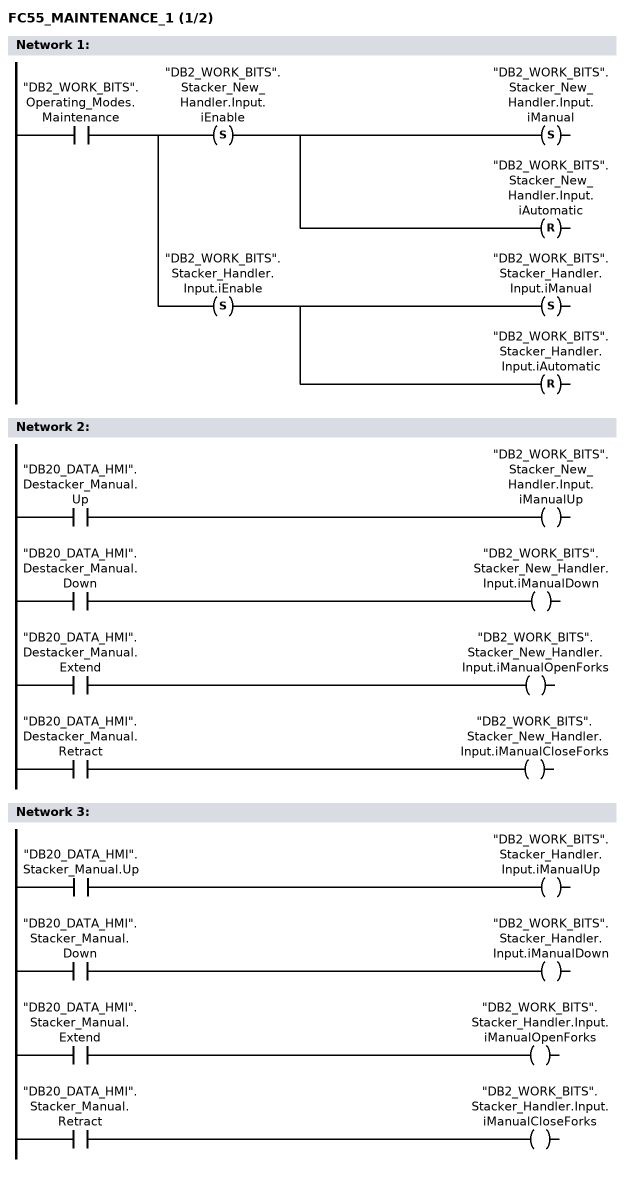
   RUNG wire#powerrail
      Contact( "DB2_WORK_BITS".Operating_Modes.Maintenance )
      wire#w1
      S_Coil( "DB2_WORK_BITS".Stacker_New_Handler.Input.iEnable )
      wire#w2
      S_Coil( "DB2_WORK_BITS".Stacker_New_Handler.Input.iManual )
   END_RUNG
   RUNG wire#w2
      R_Coil( "DB2_WORK_BITS".Stacker_New_Handler.Input.iAutomatic )
   END_RUNG
   RUNG wire#w1
      S_Coil( "DB2_WORK_BITS".Stacker_Handler.Input.iEnable )
      wire#w3
      S_Coil( "DB2_WORK_BITS".Stacker_Handler.Input.iManual )
   END_RUNG
   RUNG wire#w3
      R_Coil( "DB2_WORK_BITS".Stacker_Handler.Input.iAutomatic )
   END_RUNG
   // the same network as SCL:
   IF "DB2_WORK_BITS".Operating_Modes.Maintenance THEN
       "DB2_WORK_BITS".Stacker_New_Handler.Input.iEnable := TRUE;
       "DB2_WORK_BITS".Stacker_New_Handler.Input.iManual := TRUE;
       "DB2_WORK_BITS".Stacker_New_Handler.Input.iAutomatic := FALSE;
       "DB2_WORK_BITS".Stacker_Handler.Input.iEnable := TRUE;
       "DB2_WORK_BITS".Stacker_Handler.Input.iManual := TRUE;
       "DB2_WORK_BITS".Stacker_Handler.Input.iAutomatic := FALSE;
   END_IF;
END_REGION

REGION Network 2
   RUNG wire#powerrail
      Contact( "DB20_DATA_HMI".Destacker_Manual.Up )
      Coil( "DB2_WORK_BITS".Stacker_New_Handler.Input.iManualUp )
   END_RUNG
   RUNG wire#powerrail
      Contact( "DB20_DATA_HMI".Destacker_Manual.Down )
      Coil( "DB2_WORK_BITS".Stacker_New_Handler.Input.iManualDown )
   END_RUNG
   RUNG wire#powerrail
      Contact( "DB20_DATA_HMI".Destacker_Manual.Extend )
      Coil( "DB2_WORK_BITS".Stacker_New_Handler.Input.iManualOpenForks )
   END_RUNG
   RUNG wire#powerrail
      Contact( "DB20_DATA_HMI".Destacker_Manual.Retract )
      Coil( "DB2_WORK_BITS".Stacker_New_Handler.Input.iManualCloseForks )
   END_RUNG
   // the same network as SCL:
   "DB2_WORK_BITS".Stacker_New_Handler.Input.iManualUp := "DB20_DATA_HMI".Destacker_Manual.Up;
   "DB2_WORK_BITS".Stacker_New_Handler.Input.iManualDown := "DB20_DATA_HMI".Destacker_Manual.Down;
   "DB2_WORK_BITS".Stacker_New_Handler.Input.iManualOpenForks := "DB20_DATA_HMI".Destacker_Manual.Extend;
   "DB2_WORK_BITS".Stacker_New_Handler.Input.iManualCloseForks := "DB20_DATA_HMI".Destacker_Manual.Retract;
END_REGION

REGION Network 3
   RUNG wire#powerrail
      Contact( "DB20_DATA_HMI".Stacker_Manual.Up )
      Coil( "DB2_WORK_BITS".Stacker_Handler.Input.iManualUp )
   END_RUNG
   RUNG wire#powerrail
      Contact( "DB20_DATA_HMI".Stacker_Manual.Down )
      Coil( "DB2_WORK_BITS".Stacker_Handler.Input.iManualDown )
   END_RUNG
   RUNG wire#powerrail
      Contact( "DB20_DATA_HMI".Stacker_Manual.Extend )
      Coil( "DB2_WORK_BITS".Stacker_Handler.Input.iManualOpenForks )
   END_RUNG
   RUNG wire#powerrail
      Contact( "DB20_DATA_HMI".Stacker_Manual.Retract )
      Coil( "DB2_WORK_BITS".Stacker_Handler.Input.iManualCloseForks )
   END_RUNG
   // the same network as SCL:
   "DB2_WORK_BITS".Stacker_Handler.Input.iManualUp := "DB20_DATA_HMI".Stacker_Manual.Up;
   "DB2_WORK_BITS".Stacker_Handler.Input.iManualDown := "DB20_DATA_HMI".Stacker_Manual.Down;
   "DB2_WORK_BITS".Stacker_Handler.Input.iManualOpenForks := "DB20_DATA_HMI".Stacker_Manual.Extend;
   "DB2_WORK_BITS".Stacker_Handler.Input.iManualCloseForks := "DB20_DATA_HMI".Stacker_Manual.Retract;
END_REGION

REGION Network 4
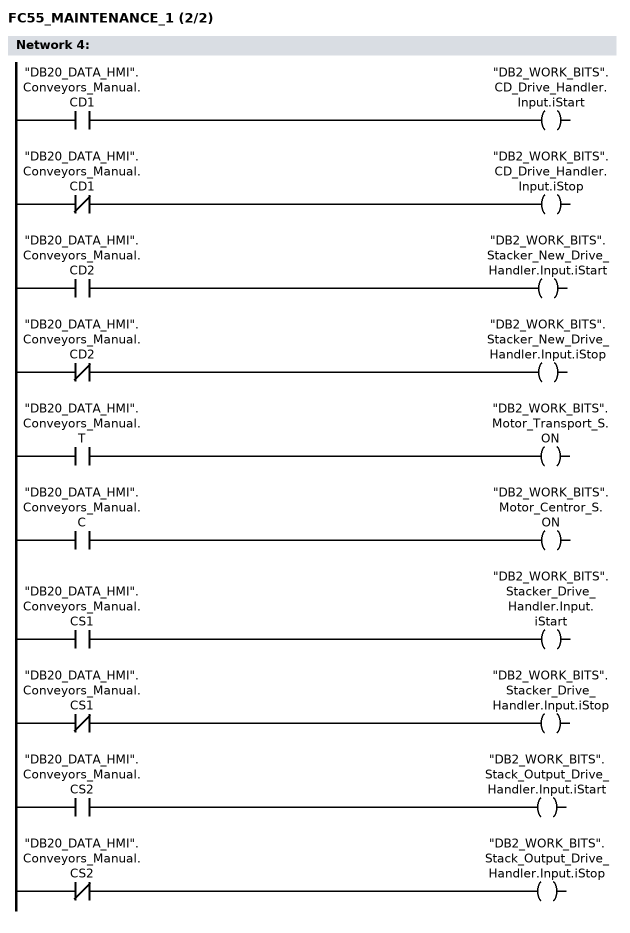
   RUNG wire#powerrail
      Contact( "DB20_DATA_HMI".Conveyors_Manual.CD1 )
      Coil( "DB2_WORK_BITS".CD_Drive_Handler.Input.iStart )
   END_RUNG
   RUNG wire#powerrail
      I_Contact( "DB20_DATA_HMI".Conveyors_Manual.CD1 )
      Coil( "DB2_WORK_BITS".CD_Drive_Handler.Input.iStop )
   END_RUNG
   RUNG wire#powerrail
      Contact( "DB20_DATA_HMI".Conveyors_Manual.CD2 )
      Coil( "DB2_WORK_BITS".Stacker_New_Drive_Handler.Input.iStart )
   END_RUNG
   RUNG wire#powerrail
      I_Contact( "DB20_DATA_HMI".Conveyors_Manual.CD2 )
      Coil( "DB2_WORK_BITS".Stacker_New_Drive_Handler.Input.iStop )
   END_RUNG
   RUNG wire#powerrail
      Contact( "DB20_DATA_HMI".Conveyors_Manual.T )
      Coil( "DB2_WORK_BITS".Motor_Transport_S.ON )
   END_RUNG
   RUNG wire#powerrail
      Contact( "DB20_DATA_HMI".Conveyors_Manual.C )
      Coil( "DB2_WORK_BITS".Motor_Centror_S.ON )
   END_RUNG
   RUNG wire#powerrail
      Contact( "DB20_DATA_HMI".Conveyors_Manual.CS1 )
      Coil( "DB2_WORK_BITS".Stacker_Drive_Handler.Input.iStart )
   END_RUNG
   RUNG wire#powerrail
      I_Contact( "DB20_DATA_HMI".Conveyors_Manual.CS1 )
      Coil( "DB2_WORK_BITS".Stacker_Drive_Handler.Input.iStop )
   END_RUNG
   RUNG wire#powerrail
      Contact( "DB20_DATA_HMI".Conveyors_Manual.CS2 )
      Coil( "DB2_WORK_BITS".Stack_Output_Drive_Handler.Input.iStart )
   END_RUNG
   RUNG wire#powerrail
      I_Contact( "DB20_DATA_HMI".Conveyors_Manual.CS2 )
      Coil( "DB2_WORK_BITS".Stack_Output_Drive_Handler.Input.iStop )
   END_RUNG
   // the same network as SCL:
   "DB2_WORK_BITS".CD_Drive_Handler.Input.iStart := "DB20_DATA_HMI".Conveyors_Manual.CD1;
   "DB2_WORK_BITS".CD_Drive_Handler.Input.iStop := NOT "DB20_DATA_HMI".Conveyors_Manual.CD1;
   "DB2_WORK_BITS".Stacker_New_Drive_Handler.Input.iStart := "DB20_DATA_HMI".Conveyors_Manual.CD2;
   "DB2_WORK_BITS".Stacker_New_Drive_Handler.Input.iStop := NOT "DB20_DATA_HMI".Conveyors_Manual.CD2;
   "DB2_WORK_BITS".Motor_Transport_S.ON := "DB20_DATA_HMI".Conveyors_Manual.T;
   "DB2_WORK_BITS".Motor_Centror_S.ON := "DB20_DATA_HMI".Conveyors_Manual.C;
   "DB2_WORK_BITS".Stacker_Drive_Handler.Input.iStart := "DB20_DATA_HMI".Conveyors_Manual.CS1;
   "DB2_WORK_BITS".Stacker_Drive_Handler.Input.iStop := NOT "DB20_DATA_HMI".Conveyors_Manual.CS1;
   "DB2_WORK_BITS".Stack_Output_Drive_Handler.Input.iStart := "DB20_DATA_HMI".Conveyors_Manual.CS2;
   "DB2_WORK_BITS".Stack_Output_Drive_Handler.Input.iStop := NOT "DB20_DATA_HMI".Conveyors_Manual.CS2;
END_REGION
END_FUNCTION

FUNCTION "FC58_SAFETY" : Void   // FC58, LAD
{ S7_Optimized_Access := 'TRUE' }
VERSION : 0.1
BEGIN

REGION Network 1: Stacker
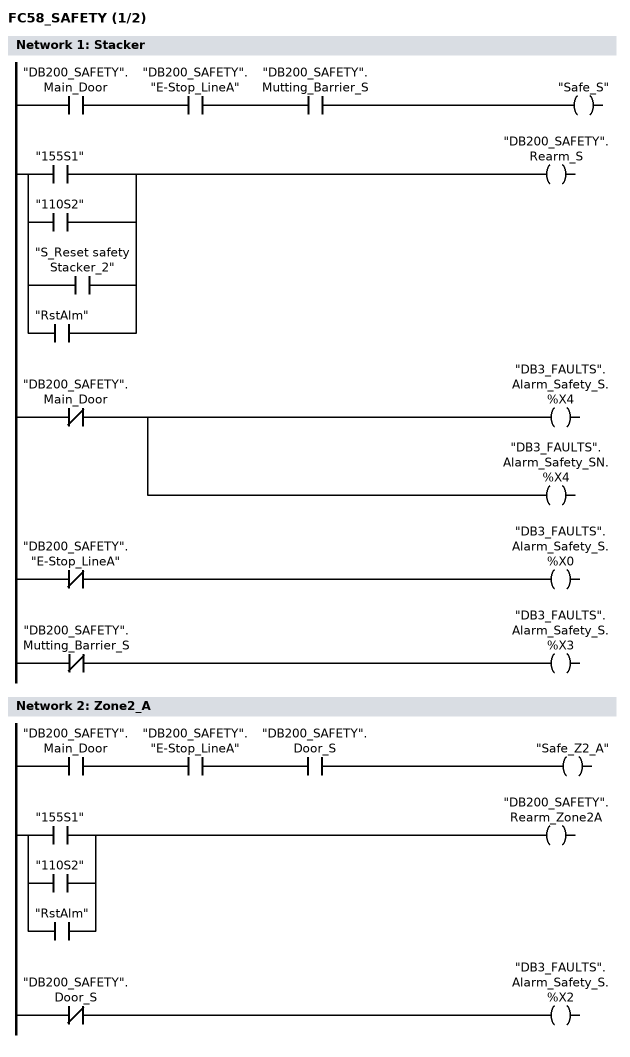
   RUNG wire#powerrail
      Contact( "DB200_SAFETY".Main_Door )
      Contact( "DB200_SAFETY"."E-Stop_LineA" )
      Contact( "DB200_SAFETY".Mutting_Barrier_S )
      Coil( "Safe_S" )
   END_RUNG
   RUNG wire#powerrail
      Contact( "155S1" )
      wire#w1
      Coil( "DB200_SAFETY".Rearm_S )
   END_RUNG
   RUNG wire#powerrail
      Contact( "110S2" )
   END_RUNG wire#w1
   RUNG wire#powerrail
      Contact( "S_Reset safety Stacker_2" )
   END_RUNG wire#w1
   RUNG wire#powerrail
      Contact( "RstAlm" )
   END_RUNG wire#w1
   RUNG wire#powerrail
      I_Contact( "DB200_SAFETY".Main_Door )
      wire#w2
      Coil( "DB3_FAULTS".Alarm_Safety_S.%X4 )
   END_RUNG
   RUNG wire#w2
      Coil( "DB3_FAULTS".Alarm_Safety_SN.%X4 )
   END_RUNG
   RUNG wire#powerrail
      I_Contact( "DB200_SAFETY"."E-Stop_LineA" )
      Coil( "DB3_FAULTS".Alarm_Safety_S.%X0 )
   END_RUNG
   RUNG wire#powerrail
      I_Contact( "DB200_SAFETY".Mutting_Barrier_S )
      Coil( "DB3_FAULTS".Alarm_Safety_S.%X3 )
   END_RUNG
   // the same network as SCL:
   "Safe_S" := "DB200_SAFETY".Main_Door AND "DB200_SAFETY"."E-Stop_LineA" AND "DB200_SAFETY".Mutting_Barrier_S;
   "DB200_SAFETY".Rearm_S := "155S1" OR "110S2" OR "S_Reset safety Stacker_2" OR "RstAlm";
   "DB3_FAULTS".Alarm_Safety_S.%X4 := NOT "DB200_SAFETY".Main_Door;
   "DB3_FAULTS".Alarm_Safety_SN.%X4 := NOT "DB200_SAFETY".Main_Door;
   "DB3_FAULTS".Alarm_Safety_S.%X0 := NOT "DB200_SAFETY"."E-Stop_LineA";
   "DB3_FAULTS".Alarm_Safety_S.%X3 := NOT "DB200_SAFETY".Mutting_Barrier_S;
END_REGION

REGION Network 2: Zone2_A
   RUNG wire#powerrail
      Contact( "DB200_SAFETY".Main_Door )
      Contact( "DB200_SAFETY"."E-Stop_LineA" )
      Contact( "DB200_SAFETY".Door_S )
      Coil( "Safe_Z2_A" )
   END_RUNG
   RUNG wire#powerrail
      Contact( "155S1" )
      wire#w1
      Coil( "DB200_SAFETY".Rearm_Zone2A )
   END_RUNG
   RUNG wire#powerrail
      Contact( "110S2" )
   END_RUNG wire#w1
   RUNG wire#powerrail
      Contact( "RstAlm" )
   END_RUNG wire#w1
   RUNG wire#powerrail
      I_Contact( "DB200_SAFETY".Door_S )
      Coil( "DB3_FAULTS".Alarm_Safety_S.%X2 )
   END_RUNG
   // the same network as SCL:
   "Safe_Z2_A" := "DB200_SAFETY".Main_Door AND "DB200_SAFETY"."E-Stop_LineA" AND "DB200_SAFETY".Door_S;
   "DB200_SAFETY".Rearm_Zone2A := "155S1" OR "110S2" OR "RstAlm";
   "DB3_FAULTS".Alarm_Safety_S.%X2 := NOT "DB200_SAFETY".Door_S;
END_REGION

REGION Network 3: Stacker_New
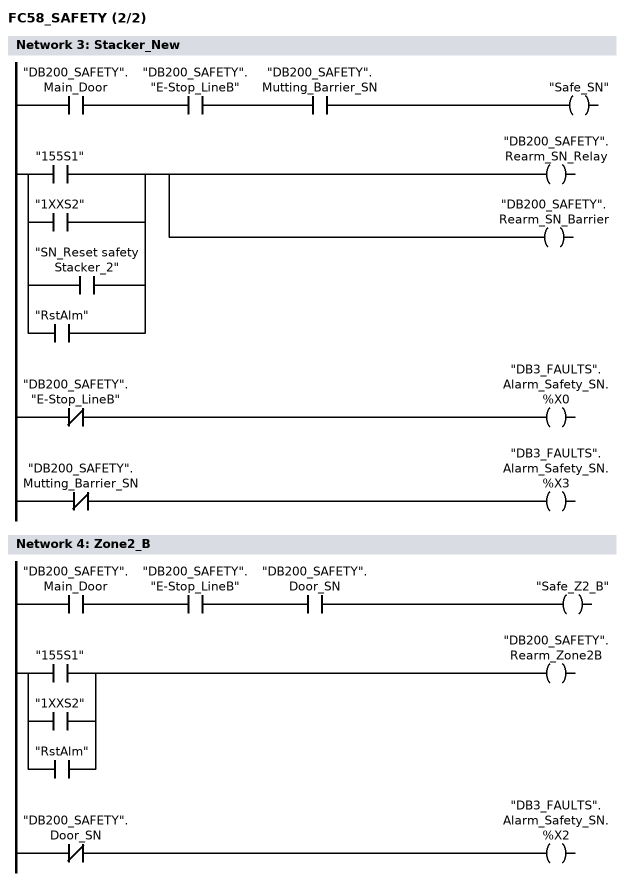
   RUNG wire#powerrail
      Contact( "DB200_SAFETY".Main_Door )
      Contact( "DB200_SAFETY"."E-Stop_LineB" )
      Contact( "DB200_SAFETY".Mutting_Barrier_SN )
      Coil( "Safe_SN" )
   END_RUNG
   RUNG wire#powerrail
      Contact( "155S1" )
      wire#w1
      Coil( "DB200_SAFETY".Rearm_SN_Relay )
   END_RUNG
   RUNG wire#powerrail
      Contact( "1XXS2" )
   END_RUNG wire#w1
   RUNG wire#powerrail
      Contact( "SN_Reset safety Stacker_2" )
   END_RUNG wire#w1
   RUNG wire#powerrail
      Contact( "RstAlm" )
   END_RUNG wire#w1
   RUNG wire#w1
      Coil( "DB200_SAFETY".Rearm_SN_Barrier )
   END_RUNG
   RUNG wire#powerrail
      I_Contact( "DB200_SAFETY"."E-Stop_LineB" )
      Coil( "DB3_FAULTS".Alarm_Safety_SN.%X0 )
   END_RUNG
   RUNG wire#powerrail
      I_Contact( "DB200_SAFETY".Mutting_Barrier_SN )
      Coil( "DB3_FAULTS".Alarm_Safety_SN.%X3 )
   END_RUNG
   // the same network as SCL:
   "Safe_SN" := "DB200_SAFETY".Main_Door AND "DB200_SAFETY"."E-Stop_LineB" AND "DB200_SAFETY".Mutting_Barrier_SN;
   "DB200_SAFETY".Rearm_SN_Relay := "155S1" OR "1XXS2" OR "SN_Reset safety Stacker_2" OR "RstAlm";
   "DB200_SAFETY".Rearm_SN_Barrier := "DB200_SAFETY".Rearm_SN_Relay;
   "DB3_FAULTS".Alarm_Safety_SN.%X0 := NOT "DB200_SAFETY"."E-Stop_LineB";
   "DB3_FAULTS".Alarm_Safety_SN.%X3 := NOT "DB200_SAFETY".Mutting_Barrier_SN;
END_REGION

REGION Network 4: Zone2_B
   RUNG wire#powerrail
      Contact( "DB200_SAFETY".Main_Door )
      Contact( "DB200_SAFETY"."E-Stop_LineB" )
      Contact( "DB200_SAFETY".Door_SN )
      Coil( "Safe_Z2_B" )
   END_RUNG
   RUNG wire#powerrail
      Contact( "155S1" )
      wire#w1
      Coil( "DB200_SAFETY".Rearm_Zone2B )
   END_RUNG
   RUNG wire#powerrail
      Contact( "1XXS2" )
   END_RUNG wire#w1
   RUNG wire#powerrail
      Contact( "RstAlm" )
   END_RUNG wire#w1
   RUNG wire#powerrail
      I_Contact( "DB200_SAFETY".Door_SN )
      Coil( "DB3_FAULTS".Alarm_Safety_SN.%X2 )
   END_RUNG
   // the same network as SCL:
   "Safe_Z2_B" := "DB200_SAFETY".Main_Door AND "DB200_SAFETY"."E-Stop_LineB" AND "DB200_SAFETY".Door_SN;
   "DB200_SAFETY".Rearm_Zone2B := "155S1" OR "1XXS2" OR "RstAlm";
   "DB3_FAULTS".Alarm_Safety_SN.%X2 := NOT "DB200_SAFETY".Door_SN;
END_REGION
END_FUNCTION

FUNCTION "FC100_CountDaily" : Void   // FC100, SCL
{ S7_Optimized_Access := 'TRUE' }
VERSION : 0.1
   VAR_INPUT
      SignalToCount : Bool;
      Reset : Bool;
   END_VAR
   VAR_IN_OUT
      CurrentValue : UDInt;
   END_VAR
   VAR_TEMP
      timeofday : DTL;
      ret : Int;
   END_VAR
BEGIN
   #ret := RD_LOC_T(#timeofday);
END_FUNCTION

ORGANIZATION_BLOCK "Main"   // OB1, LAD, ProgramCycle
TITLE = "Main Program Sweep (Cycle)"
{ S7_Optimized_Access := 'TRUE' }
VERSION : 0.1
   VAR_INPUT
      Initial_Call : Bool;   // Initial call of this OB
      Remanence : Bool;   // =True, if remanent data are available
   END_VAR
   VAR_TEMP
      Move_Block_Diag : Int;
   END_VAR
BEGIN

REGION Network 1
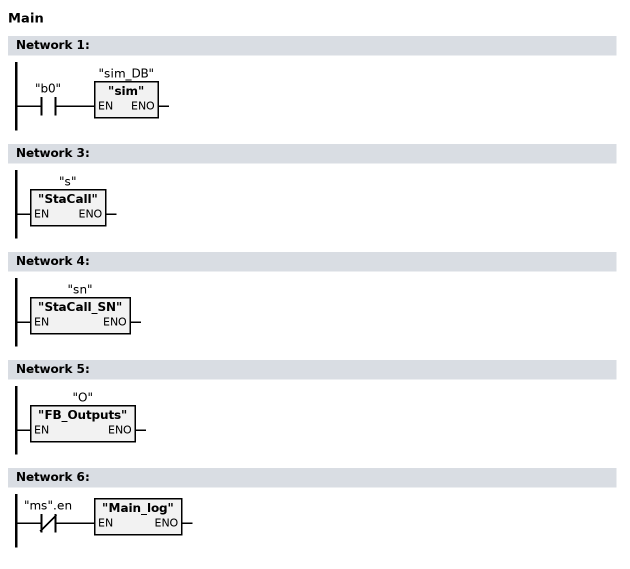
   RUNG wire#powerrail
      Contact( "b0" )
      "sim_DB"()
   END_RUNG
   // the same network as SCL:
   IF "b0" THEN
       "sim_DB"();   // "sim"
   END_IF;
END_REGION

REGION Network 2 (SCL)
   "FC58_SAFETY"();
   "FC6_OUTPUTS"();

   "FC60_MappingIn"();

   "FC3_FAULTS"();
   "FB_GEN_DB"();

   "FC_AckOpTranzit"();


   "FC52_STACKING"();
   "FC52_STACKING_New"();

   //"FC55_MAINTENANCE"();
   "FC20_HMI"();
   "FB_IntervalTrigger_DB"();
   "FB_EnergyCounter_DB"(ibMeterPulse := "DB2_WORK_BITS".Consumption_Pulse,
                         ibHourChange := "FB_IntervalTrigger_DB".bHourChanged,
                        ibDayChange := "FB_IntervalTrigger_DB".bDayChanged,
                         ibMonthChange := "FB_IntervalTrigger_DB".bMonthChanged,
                         ibReset := FALSE);
   "FB_AlarmCounter_DB"();
   "FB_ProductionStatistics_DB"(ibDestroy:="DB2_WORK_BITS".SQ_Outfeed_Stack_SN,
                                ibRepair:="DB2_WORK_BITS".Transport_Conveyor_SQs.SQ_Repaired_Pallet[0] OR "DB2_WORK_BITS".Transport_Conveyor_SQs.SQ_Repaired_Pallet[1],
                                ibDayChange:="FB_IntervalTrigger_DB".bDayChanged,
                                ibMonthChange:="FB_IntervalTrigger_DB".bMonthChanged);
END_REGION

REGION Network 3
   RUNG wire#powerrail
      "s"()
   END_RUNG
   // the same network as SCL:
   "s"();   // "StaCall"
END_REGION

REGION Network 4
   RUNG wire#powerrail
      "sn"()
   END_RUNG
   // the same network as SCL:
   "sn"();   // "StaCall_SN"
END_REGION

REGION Network 5
   RUNG wire#powerrail
      "O"()
   END_RUNG
   // the same network as SCL:
   "O"();   // "FB_Outputs"
END_REGION

REGION Network 6
   RUNG wire#powerrail
      I_Contact( "ms".en )
      "Main_log"()
   END_RUNG
   // the same network as SCL:
   IF NOT "ms".en THEN "Main_log"(); END_IF;
END_REGION
END_ORGANIZATION_BLOCK

ORGANIZATION_BLOCK "OB82_I/O_FLT"   // OB82, LAD, DiagnosticErrorInterrupt
{ S7_Optimized_Access := 'TRUE' }
VERSION : 0.1
   VAR_INPUT
      IO_State : Word;   // IO state of the HW object
      LADDR : Hw_Any;   // Hardware identifier
      Channel : UInt;   // Channel number
      MultiError : Bool;   // =true if more than one error is present
   END_VAR
BEGIN
END_ORGANIZATION_BLOCK

ORGANIZATION_BLOCK "OB100_COMPLETE_RESTART"   // OB100, LAD, Startup
TITLE = "Complete Restart"
{ S7_Optimized_Access := 'TRUE' }
VERSION : 0.1
   VAR_INPUT
      LostRetentive : Bool;   // True if retentive data are lost
      LostRTC : Bool;   // True if date and time are lost
   END_VAR
BEGIN
END_ORGANIZATION_BLOCK

// folder: Stacker_New

FUNCTION_BLOCK "StaCall_SN"   // FB15, LAD
{ S7_Optimized_Access := 'TRUE' }
VERSION : 0.1
   VAR
      f : Array[0..10] of "sta_SN";
      tranzit : Array[0..10] of Bool;
      Range_LS_1 : Bool;
      Range_LS_2 : Bool;
      Range_LS_3 : Bool;
      PrezPalStackLength : Bool;
      PrezPalStackAnyLength : Bool;
      PrezPalStackAny : Bool;
      DeliveryStack : Bool;
      StivStat : USInt;
      nAc : USInt;
      tmrSnzCentr : TON_TIME;
      tmr : Array[0..8] of IEC_TIMER;
   END_VAR
   VAR_TEMP
      to_ce : Bool;
      to_cm : Bool;
      cmdLiftUpO : Bool;
      tranzit12 : Bool;
   END_VAR
   VAR CONSTANT
      _nop0 : Int := 0;
      _op1 : Int := 1;
      _cen : Int := 3;
      _stack : Int := 4;
      _evac : Int := 5;
      _nop : Int := 6;
   END_VAR
   VAR_TEMP   // added for the SCL form of the ladder/FBD networks
      _w1 : Bool;
      _w2 : Bool;
      _w3 : Bool;
   END_VAR
BEGIN

REGION Network 1: Force init
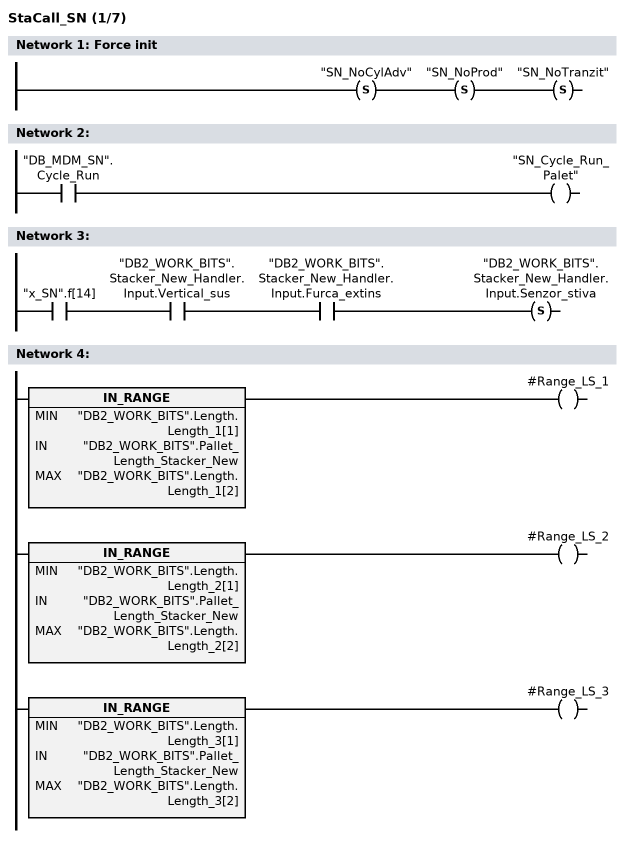
   RUNG wire#powerrail
      S_Coil( "SN_NoCylAdv" )
      S_Coil( "SN_NoProd" )
      S_Coil( "SN_NoTranzit" )
   END_RUNG
   // the same network as SCL:
   "SN_NoCylAdv" := TRUE;
   "SN_NoProd" := TRUE;
   "SN_NoTranzit" := TRUE;
END_REGION

REGION Network 2
   RUNG wire#powerrail
      Contact( "DB_MDM_SN".Cycle_Run )
      Coil( "SN_Cycle_Run_Palet" )
   END_RUNG
   // the same network as SCL:
   "SN_Cycle_Run_Palet" := "DB_MDM_SN".Cycle_Run;
END_REGION

REGION Network 3
   RUNG wire#powerrail
      Contact( "x_SN".f[14] )
      Contact( "DB2_WORK_BITS".Stacker_New_Handler.Input.Vertical_sus )
      Contact( "DB2_WORK_BITS".Stacker_New_Handler.Input.Furca_extins )
      S_Coil( "DB2_WORK_BITS".Stacker_New_Handler.Input.Senzor_stiva )
   END_RUNG
   // the same network as SCL:
   IF "x_SN".f[14] AND "DB2_WORK_BITS".Stacker_New_Handler.Input.Vertical_sus AND "DB2_WORK_BITS".Stacker_New_Handler.Input.Furca_extins THEN
       "DB2_WORK_BITS".Stacker_New_Handler.Input.Senzor_stiva := TRUE;
   END_IF;
END_REGION

REGION Network 4
   RUNG wire#powerrail
      { S7_Templates := "SrcType := Int" } InRange(min := "DB2_WORK_BITS".Length.Length_1[1], in := "DB2_WORK_BITS".Pallet_Length_Stacker_New, max := "DB2_WORK_BITS".Length.Length_1[2])
      Coil( #Range_LS_1 )
   END_RUNG
   RUNG wire#powerrail
      { S7_Templates := "SrcType := Int" } InRange(min := "DB2_WORK_BITS".Length.Length_2[1], in := "DB2_WORK_BITS".Pallet_Length_Stacker_New, max := "DB2_WORK_BITS".Length.Length_2[2])
      Coil( #Range_LS_2 )
   END_RUNG
   RUNG wire#powerrail
      { S7_Templates := "SrcType := Int" } InRange(min := "DB2_WORK_BITS".Length.Length_3[1], in := "DB2_WORK_BITS".Pallet_Length_Stacker_New, max := "DB2_WORK_BITS".Length.Length_3[2])
      Coil( #Range_LS_3 )
   END_RUNG
   // the same network as SCL:
   #Range_LS_1 := ("DB2_WORK_BITS".Length.Length_1[1] <= "DB2_WORK_BITS".Pallet_Length_Stacker_New) AND ("DB2_WORK_BITS".Pallet_Length_Stacker_New <= "DB2_WORK_BITS".Length.Length_1[2]);
   #Range_LS_2 := ("DB2_WORK_BITS".Length.Length_2[1] <= "DB2_WORK_BITS".Pallet_Length_Stacker_New) AND ("DB2_WORK_BITS".Pallet_Length_Stacker_New <= "DB2_WORK_BITS".Length.Length_2[2]);
   #Range_LS_3 := ("DB2_WORK_BITS".Length.Length_3[1] <= "DB2_WORK_BITS".Pallet_Length_Stacker_New) AND ("DB2_WORK_BITS".Pallet_Length_Stacker_New <= "DB2_WORK_BITS".Length.Length_3[2]);
END_REGION

REGION Network 5: 1 Op1- - Reparare palete Zona B
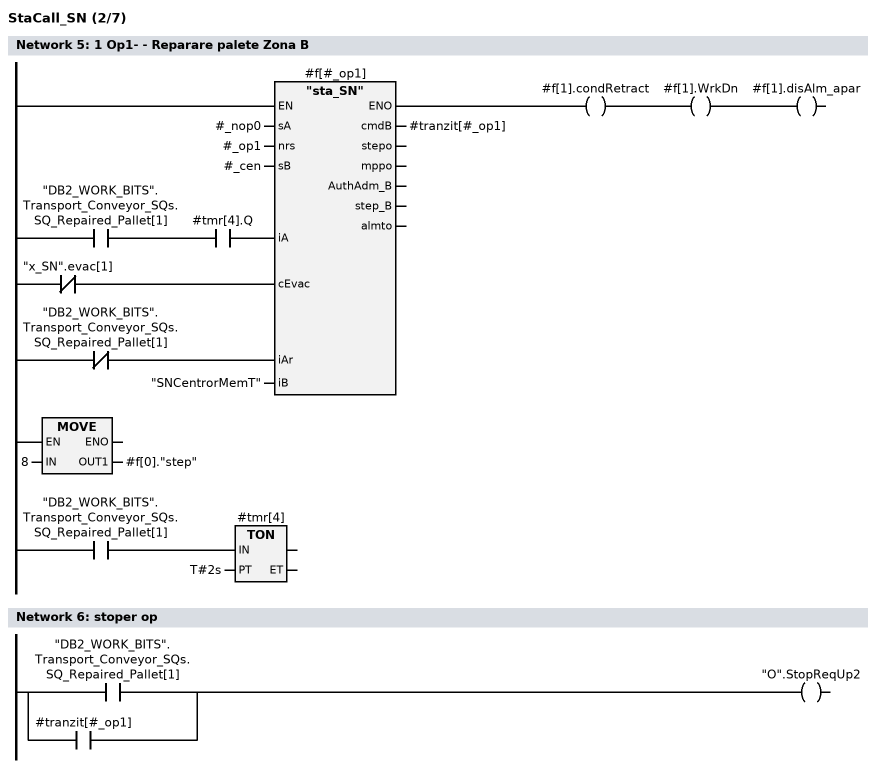
   #f[#_op1](sA := #_nop0,   // "sta_SN"
             nrs := #_op1,
             sB := #_cen,
             iA := "DB2_WORK_BITS".Transport_Conveyor_SQs.SQ_Repaired_Pallet[1] AND #tmr[4].Q,
             cEvac := NOT "x_SN".evac[1],
             iAr := NOT "DB2_WORK_BITS".Transport_Conveyor_SQs.SQ_Repaired_Pallet[1],
             iB := "SNCentrorMemT",
             cmdB => #tranzit[#_op1],
             ENO => #_w1);
   #f[1].condRetract := #_w1;
   #f[1].WrkDn := #_w1;
   #f[1].disAlm_apar := #_w1;
   #f[0]."step" := 8;
   #tmr[4].TON(IN := "DB2_WORK_BITS".Transport_Conveyor_SQs.SQ_Repaired_Pallet[1], PT := T#2s);
END_REGION

REGION Network 6: stoper op
   RUNG wire#powerrail
      Contact( "DB2_WORK_BITS".Transport_Conveyor_SQs.SQ_Repaired_Pallet[1] )
      wire#w1
      Coil( "O".StopReqUp2 )
   END_RUNG
   RUNG wire#powerrail
      Contact( #tranzit[#_op1] )
   END_RUNG wire#w1
   // the same network as SCL:
   "O".StopReqUp2 := "DB2_WORK_BITS".Transport_Conveyor_SQs.SQ_Repaired_Pallet[1] OR #tranzit[#_op1];
END_REGION

REGION Network 7
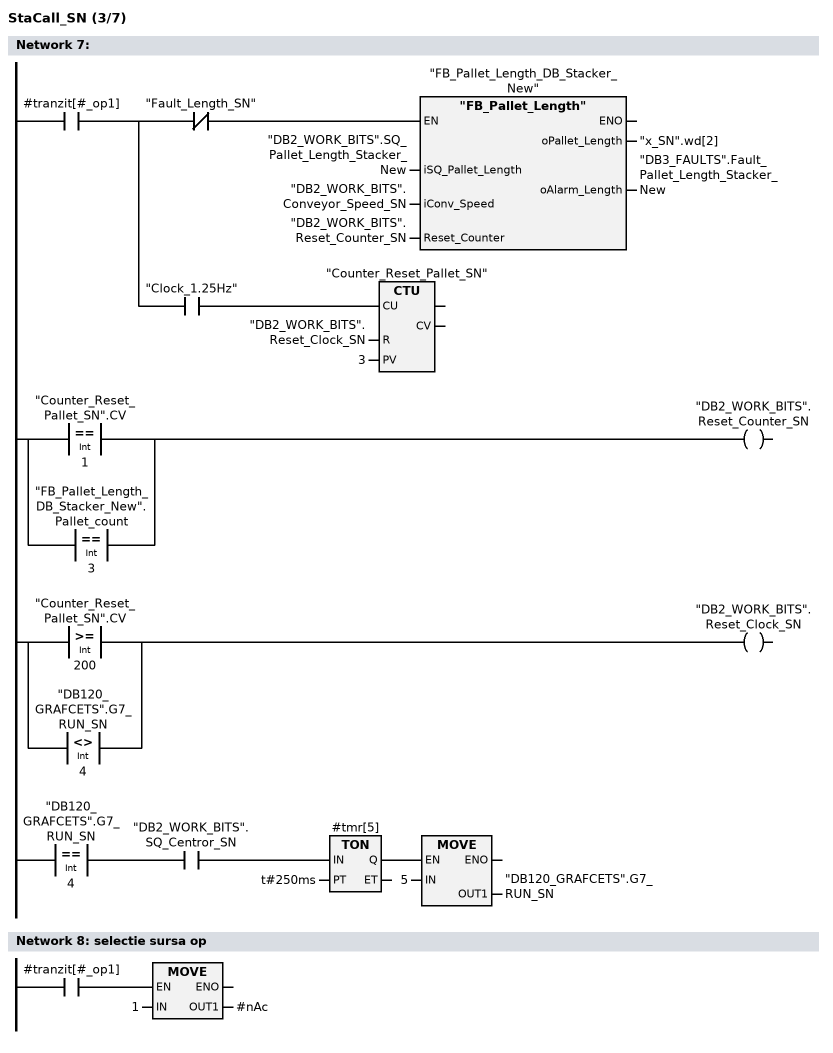
   IF #tranzit[#_op1] AND NOT "Fault_Length_SN" THEN
       "FB_Pallet_Length_DB_Stacker_New"(iSQ_Pallet_Length := "DB2_WORK_BITS".SQ_Pallet_Length_Stacker_New,   // "FB_Pallet_Length"
                               iConv_Speed := "DB2_WORK_BITS".Conveyor_Speed_SN,
                               Reset_Counter := "DB2_WORK_BITS".Reset_Counter_SN,
                               oPallet_Length => "x_SN".wd[2],
                               oAlarm_Length => "DB3_FAULTS".Fault_Pallet_Length_Stacker_New);
   END_IF;
   "Counter_Reset_Pallet_SN".CTU(CU := #tranzit[#_op1] AND "Clock_1.25Hz",
                           R := "DB2_WORK_BITS".Reset_Clock_SN,
                           PV := 3);
   "DB2_WORK_BITS".Reset_Counter_SN := ("Counter_Reset_Pallet_SN".CV = 1) OR ("FB_Pallet_Length_DB_Stacker_New".Pallet_count = 3);
   "DB2_WORK_BITS".Reset_Clock_SN := ("Counter_Reset_Pallet_SN".CV >= 200) OR ("DB120_GRAFCETS".G7_RUN_SN <> 4);
   #tmr[5].TON(IN := ("DB120_GRAFCETS".G7_RUN_SN = 4) AND "DB2_WORK_BITS".SQ_Centror_SN, PT := t#250ms);
   IF #tmr[5].Q THEN "DB120_GRAFCETS".G7_RUN_SN := 5; END_IF;
END_REGION

REGION Network 8: selectie sursa op
   RUNG wire#powerrail
      Contact( #tranzit[#_op1] )
      Move(in := 1, out1 => #nAc)
   END_RUNG
   // the same network as SCL:
   IF #tranzit[#_op1] THEN #nAc := 1; END_IF;
END_REGION

REGION Network 9: senz stop stk
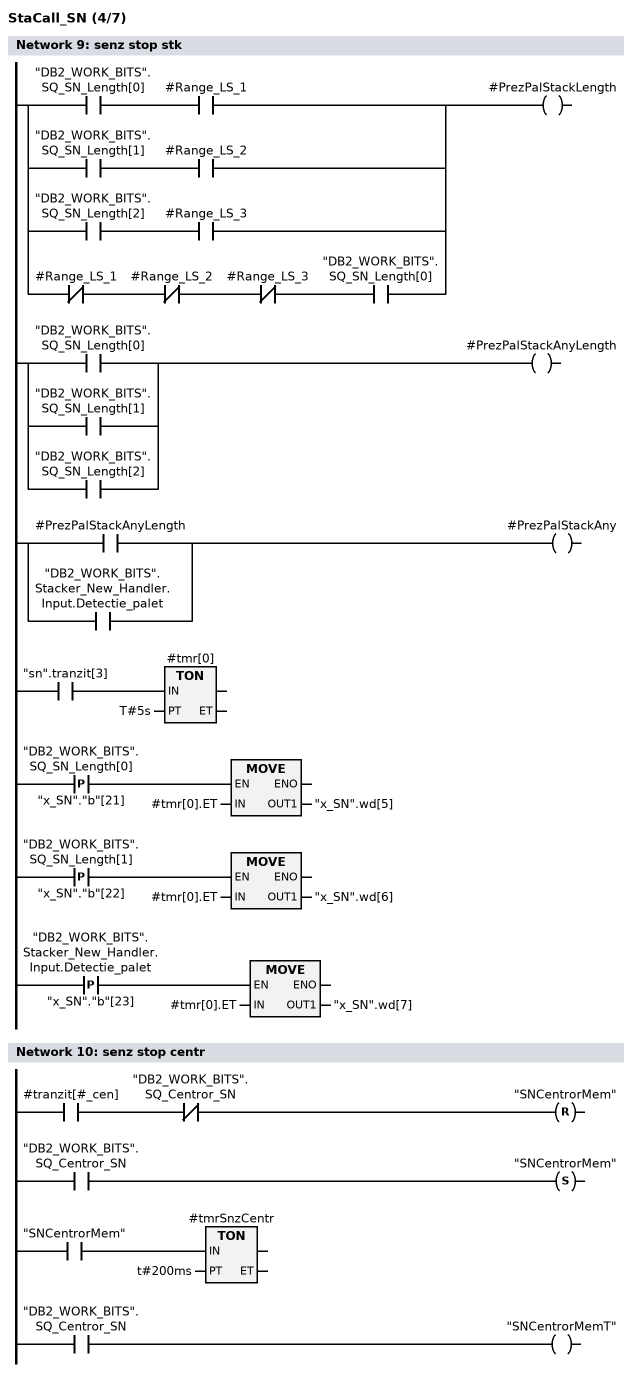
   #PrezPalStackLength := ("DB2_WORK_BITS".SQ_SN_Length[0] AND #Range_LS_1) OR ("DB2_WORK_BITS".SQ_SN_Length[1] AND #Range_LS_2) OR ("DB2_WORK_BITS".SQ_SN_Length[2] AND #Range_LS_3) OR (NOT #Range_LS_1 AND NOT #Range_LS_2 AND NOT #Range_LS_3 AND "DB2_WORK_BITS".SQ_SN_Length[0]);
   #PrezPalStackAnyLength := "DB2_WORK_BITS".SQ_SN_Length[0] OR "DB2_WORK_BITS".SQ_SN_Length[1] OR "DB2_WORK_BITS".SQ_SN_Length[2];
   #PrezPalStackAny := #PrezPalStackAnyLength OR "DB2_WORK_BITS".Stacker_New_Handler.Input.Detectie_palet;
   #tmr[0].TON(IN := "sn".tranzit[3], PT := T#5s);
   #_w1 := "DB2_WORK_BITS".SQ_SN_Length[0] AND NOT "x_SN"."b"[21];   // rising edge of "DB2_WORK_BITS".SQ_SN_Length[0]
   "x_SN"."b"[21] := "DB2_WORK_BITS".SQ_SN_Length[0];
   IF #_w1 THEN "x_SN".wd[5] := #tmr[0].ET; END_IF;
   #_w2 := "DB2_WORK_BITS".SQ_SN_Length[1] AND NOT "x_SN"."b"[22];   // rising edge of "DB2_WORK_BITS".SQ_SN_Length[1]
   "x_SN"."b"[22] := "DB2_WORK_BITS".SQ_SN_Length[1];
   IF #_w2 THEN "x_SN".wd[6] := #tmr[0].ET; END_IF;
   #_w3 := "DB2_WORK_BITS".Stacker_New_Handler.Input.Detectie_palet AND NOT "x_SN"."b"[23];   // rising edge of "DB2_WORK_BITS".Stacker_New_Handler.Input.Detectie_palet
   "x_SN"."b"[23] := "DB2_WORK_BITS".Stacker_New_Handler.Input.Detectie_palet;
   IF #_w3 THEN "x_SN".wd[7] := #tmr[0].ET; END_IF;
END_REGION

REGION Network 10: senz stop centr
   IF #tranzit[#_cen] AND NOT "DB2_WORK_BITS".SQ_Centror_SN THEN "SNCentrorMem" := FALSE; END_IF;
   IF "DB2_WORK_BITS".SQ_Centror_SN THEN "SNCentrorMem" := TRUE; END_IF;
   #tmrSnzCentr(IN := "SNCentrorMem", PT := t#200ms);   // TON
   "SNCentrorMemT" := "DB2_WORK_BITS".SQ_Centror_SN;
END_REGION

REGION Network 11: 3- Centror
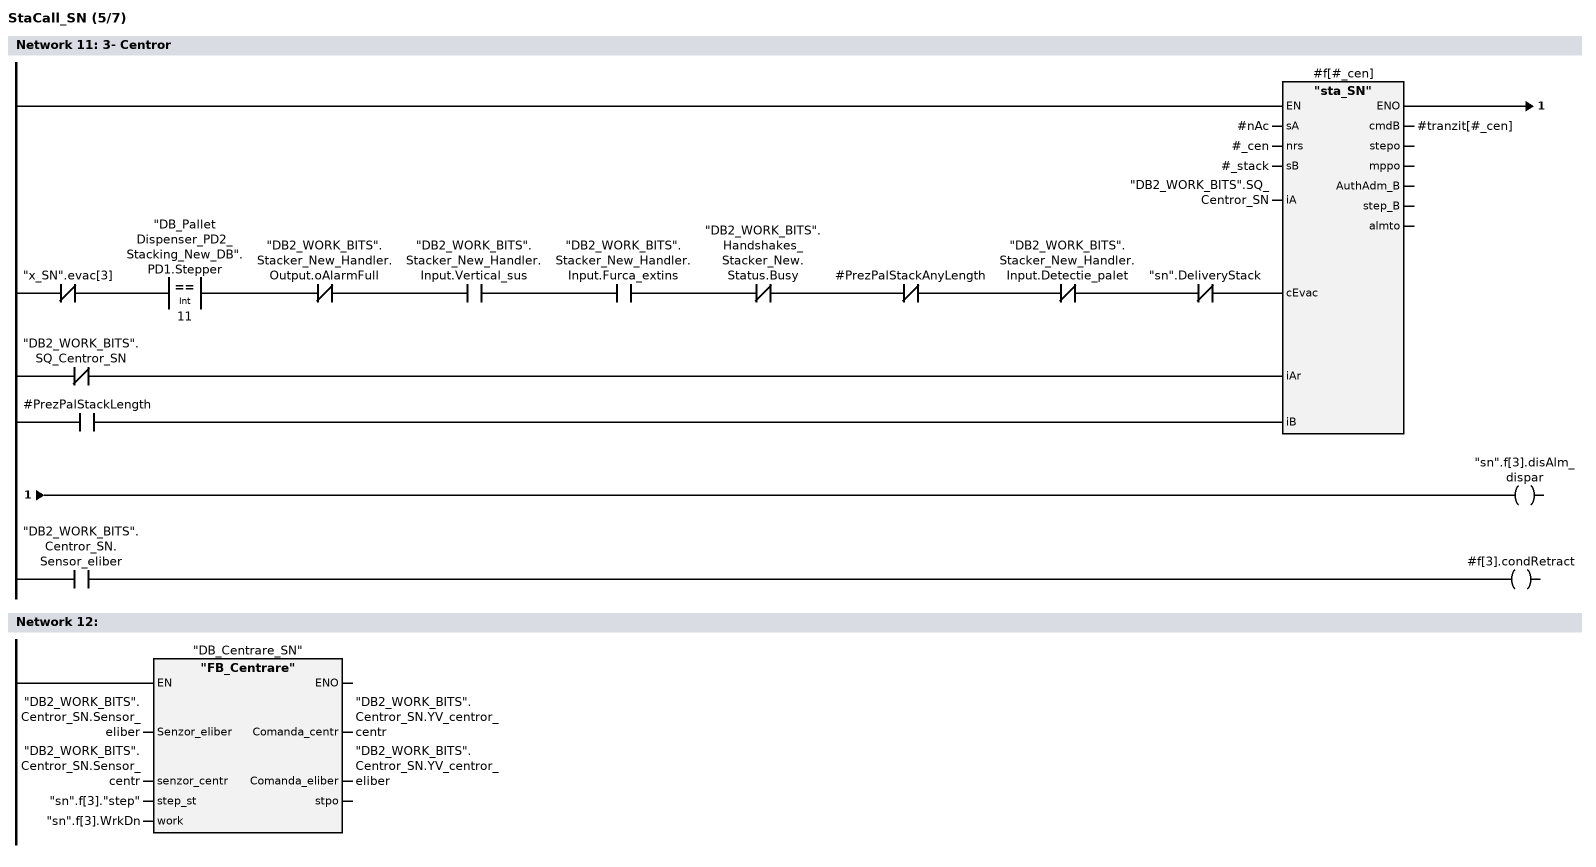
   RUNG wire#powerrail
      #f[#_cen](cEvac := wire#w1, iAr := wire#w2, iB := wire#w3, sA := #nAc, nrs := #_cen, sB := #_stack, iA := "DB2_WORK_BITS".SQ_Centror_SN, cmdB => #tranzit[#_cen], stepo =>, mppo =>, AuthAdm_B =>, step_B =>, almto =>)
      Coil( "sn".f[3].disAlm_dispar )
   END_RUNG
   RUNG wire#powerrail
      I_Contact( "x_SN".evac[3] )
      { S7_Templates := "SrcType := Int" } EQ_Contact(in1 := "DB_PalletDispenser_PD2_Stacking_New_DB".PD1.Stepper, in2 := 11)
      I_Contact( "DB2_WORK_BITS".Stacker_New_Handler.Output.oAlarmFull )
      Contact( "DB2_WORK_BITS".Stacker_New_Handler.Input.Vertical_sus )
      Contact( "DB2_WORK_BITS".Stacker_New_Handler.Input.Furca_extins )
      I_Contact( "DB2_WORK_BITS".Handshakes_Stacker_New.Status.Busy )
      I_Contact( #PrezPalStackAnyLength )
      I_Contact( "DB2_WORK_BITS".Stacker_New_Handler.Input.Detectie_palet )
      I_Contact( "sn".DeliveryStack )
   END_RUNG wire#w1
   RUNG wire#powerrail
      I_Contact( "DB2_WORK_BITS".SQ_Centror_SN )
   END_RUNG wire#w2
   RUNG wire#powerrail
      Contact( #PrezPalStackLength )
   END_RUNG wire#w3
   RUNG wire#powerrail
      Contact( "DB2_WORK_BITS".Centror_SN.Sensor_eliber )
      Coil( #f[3].condRetract )
   END_RUNG
   // the same network as SCL:
   #f[#_cen](sA := #nAc,   // "sta_SN"
             nrs := #_cen,
             sB := #_stack,
             iA := "DB2_WORK_BITS".SQ_Centror_SN,
             cEvac := NOT "x_SN".evac[3] AND ("DB_PalletDispenser_PD2_Stacking_New_DB".PD1.Stepper = 11) AND NOT "DB2_WORK_BITS".Stacker_New_Handler.Output.oAlarmFull AND "DB2_WORK_BITS".Stacker_New_Handler.Input.Vertical_sus AND "DB2_WORK_BITS".Stacker_New_Handler.Input.Furca_extins AND NOT "DB2_WORK_BITS".Handshakes_Stacker_New.Status.Busy AND NOT #PrezPalStackAnyLength AND NOT "DB2_WORK_BITS".Stacker_New_Handler.Input.Detectie_palet AND NOT "sn".DeliveryStack,
             iAr := NOT "DB2_WORK_BITS".SQ_Centror_SN,
             iB := #PrezPalStackLength,
             cmdB => #tranzit[#_cen],
             ENO => #_w1);
   "sn".f[3].disAlm_dispar := #_w1;
   #f[3].condRetract := "DB2_WORK_BITS".Centror_SN.Sensor_eliber;
END_REGION

REGION Network 12
   RUNG wire#powerrail
      "DB_Centrare_SN"(Senzor_eliber := "DB2_WORK_BITS".Centror_SN.Sensor_eliber, senzor_centr := "DB2_WORK_BITS".Centror_SN.Sensor_centr, step_st := "sn".f[3]."step", work := "sn".f[3].WrkDn, Comanda_centr => "DB2_WORK_BITS".Centror_SN.YV_centror_centr, Comanda_eliber => "DB2_WORK_BITS".Centror_SN.YV_centror_eliber, stpo =>)
   END_RUNG
   // the same network as SCL:
   "DB_Centrare_SN"(Senzor_eliber := "DB2_WORK_BITS".Centror_SN.Sensor_eliber,   // "FB_Centrare"
                    senzor_centr := "DB2_WORK_BITS".Centror_SN.Sensor_centr,
                    step_st := "sn".f[3]."step",
                    work := "sn".f[3].WrkDn,
                    Comanda_centr => "DB2_WORK_BITS".Centror_SN.YV_centror_centr,
                    Comanda_eliber => "DB2_WORK_BITS".Centror_SN.YV_centror_eliber);
END_REGION

REGION Network 13: 4- stacker
